   IOField "I/O field_9" at 378,310 size 30x20; FormatPattern 99
      ProcessValue <- "Motors_DB_M3_Wait_On_Now"
   IOField "I/O field_10" at 378,333 size 30x20; FormatPattern 99
      ProcessValue <- "Motors_DB_M3_Wait_Off_Now"
   IOField "I/O field_11" at 313,383 size 98x20; FormatPattern 9999999999
      ProcessValue <- "Motors_DB_M3_Res_h"
   Button "Button_45" at 213,384 size 90x20; TextOff 'Force'
      on Click: InvertBit("Motors_DB_M3_CMD_Force")
      Appearance <- "Motors_DB_M3_CMD_Force"

screen "Trans" 800x480, template "Main"
   TextField "Text field_2" at 210,15 size 67x22; Text 'Датчик:'
   TextField "Text field_4" at 273,15 size 94x22; Text 'Мутность 1'
   TextField "Text field_7" at 390,18 size 43x22; Text 'вход'
   TextField "Text field_8" at 390,43 size 56x22; Text 'выход'
   IOField "I/O field_1" at 452,19 size 102x26; FormatPattern s99999.99
      ProcessValue <- "AIx_DB_Trans_1_Converter_Min_In"
   IOField "I/O field_2" at 452,41 size 102x26; FormatPattern s99999.99
      ProcessValue <- "AIx_DB_Trans_1_Converter_Min_Out"
   IOField "I/O field_3" at 551,19 size 102x26; FormatPattern s99999.99
      ProcessValue <- "AIx_DB_Trans_1_Converter_Max_In"
   IOField "I/O field_4" at 551,41 size 102x26; FormatPattern s99999.99
      ProcessValue <- "AIx_DB_Trans_1_Converter_Max_Out"
   TextField "Text field_9" at 389,68 size 101x22; Text 'Фильтрация'
   TextField "Text field_10" at 390,96 size 36x22; Text 'RTD'
   Button "Button_7" at 489,71 size 20x20; TextOff 'Text'; PictureList "ok"
      on Click: InvertBit("AIx_DB_Trans_1_Use_Filter")
      ProcessValue <- "AIx_DB_Trans_1_Use_Filter"
   Button "Button_8" at 489,96 size 20x20; TextOff 'Text'; PictureList "ok"
      on Click: InvertBit("AIx_DB_Trans_1_Use_RTD")
      ProcessValue <- "AIx_DB_Trans_1_Use_RTD"
   IOField "I/O field_5" at 516,68 size 65x25; FormatPattern 999
      ProcessValue <- "AIx_DB_Trans_1_Filter_SP"
   IOField "I/O field_6" at 516,93 size 65x25; FormatPattern 999
      ProcessValue <- "AIx_DB_Trans_1_RTD_c"
   TextField "Text field_11" at 210,36 size 79x22; Text 'Поправка'
   IOField "I/O field_7" at 293,36 size 78x23; FormatPattern s999.9
      ProcessValue <- "AIx_DB_Trans_1_Calibration"
   Button "Button_9" at 396,176 size 248x28; TextOff 'Use'
      on Click: InvertBit("AIx_DB_Trans_1_CMD_Start_A")
      Appearance <- "AIx_DB_Trans_1_CMD_Start_A"
   Button "Button_10" at 213,66 size 68x28; TextOff 'Hand'
      on Click: InvertBit("AIx_DB_Trans_1_CMD_Hand")
      Appearance <- "AIx_DB_Trans_1_CMD_Hand"
   IOField "I/O field_8" at 293,66 size 78x28; FormatPattern s9999.9
      ProcessValue <- "AIx_DB_Trans_1_Result"
   TextField "Text field_12" at 436,123 size 27x22; Text 'NC'
   TextField "Text field_13" at 437,143 size 25x22; Text 'SC'
   TextField "Text field_14" at 210,125 size 27x22; Text 'HH'
   TextField "Text field_15" at 216,145 size 16x22; Text 'H'
   TextField "Text field_16" at 217,165 size 14x22; Text 'L'
   TextField "Text field_17" at 212,186 size 23x22; Text 'LL'
   IOField "I/O field_11" at 472,123 size 58x21; FormatPattern s99999
      ProcessValue <- "AIx_DB_Trans_1_SP_NC"
   IOField "I/O field_12" at 472,143 size 58x21; FormatPattern s99999
      ProcessValue <- "AIx_DB_Trans_1_SP_SC"
   IOField "I/O field_13" at 246,125 size 58x21; FormatPattern 99999
      ProcessValue <- "AIx_DB_Trans_1_SP_HH"
   IOField "I/O field_14" at 246,145 size 58x21; FormatPattern 99999
      ProcessValue <- "AIx_DB_Trans_1_SP_H"
   IOField "I/O field_15" at 246,165 size 58x21; FormatPattern s99999
      ProcessValue <- "AIx_DB_Trans_1_SP_L"
   IOField "I/O field_16" at 246,185 size 58x21; FormatPattern s99999
      ProcessValue <- "AIx_DB_Trans_1_SP_LL"
   IOField "I/O field_17" at 546,123 size 58x21; FormatPattern 999
      ProcessValue <- "AIx_DB_Trans_1_Timers_NC_SP"
   IOField "I/O field_18" at 546,143 size 58x21; FormatPattern 999
      ProcessValue <- "AIx_DB_Trans_1_Timers_SC_SP"
   IOField "I/O field_19" at 320,125 size 58x21; FormatPattern 999
      ProcessValue <- "AIx_DB_Trans_1_Timers_HH_SP"
   IOField "I/O field_20" at 320,145 size 58x21; FormatPattern 999
      ProcessValue <- "AIx_DB_Trans_1_Timers_H_SP"
   IOField "I/O field_21" at 320,165 size 58x21; FormatPattern 999
      ProcessValue <- "AIx_DB_Trans_1_Timers_L_SP"
   IOField "I/O field_22" at 320,185 size 58x21; FormatPattern 999
      ProcessValue <- "AIx_DB_Trans_1_Timers_LL_SP"
   IOField "I/O field_23" at 582,93 size 65x25; FormatPattern s99999
      ProcessValue <- "AIx_DB_Trans_1_Signal"
   TextField "Text field_18" at 210,97 size 68x22; Text 'Уставка'
   TextField "Text field_19" at 299,97 size 79x22; Text 'Время (с)'
   TextField "Text field_1" at 214,248 size 67x22; Text 'Датчик:'
   TextField "Text field_3" at 277,248 size 94x22; Text 'Мутность 2'
   TextField "Text field_5" at 394,251 size 43x22; Text 'вход'
   TextField "Text field_6" at 394,276 size 56x22; Text 'выход'
   IOField "I/O field_9" at 456,252 size 102x26; FormatPattern s99999.99
      ProcessValue <- "AIx_DB_Trans_2_Converter_Min_In"
   IOField "I/O field_10" at 456,274 size 102x26; FormatPattern s99999.99
      ProcessValue <- "AIx_DB_Trans_2_Converter_Min_Out"
   IOField "I/O field_24" at 555,252 size 102x26; FormatPattern s99999.99
      ProcessValue <- "AIx_DB_Trans_2_Converter_Max_In"
   IOField "I/O field_25" at 555,274 size 102x26; FormatPattern s99999.99
      ProcessValue <- "AIx_DB_Trans_2_Converter_Max_Out"
   TextField "Text field_20" at 393,301 size 101x22; Text 'Фильтрация'
   TextField "Text field_21" at 394,329 size 36x22; Text 'RTD'
   Button "Button_11" at 493,304 size 20x20; TextOff 'Text'; PictureList "ok"
      on Click: InvertBit("AIx_DB_Trans_2_Use_Filter")
      ProcessValue <- "AIx_DB_Trans_2_Use_Filter"
   Button "Button_12" at 493,329 size 20x20; TextOff 'Text'; PictureList "ok"
      on Click: InvertBit("AIx_DB_Trans_2_Use_RTD")
      ProcessValue <- "AIx_DB_Trans_2_Use_RTD"
   IOField "I/O field_26" at 520,301 size 65x25; FormatPattern 999
      ProcessValue <- "AIx_DB_Trans_2_Filter_SP"
   IOField "I/O field_27" at 520,326 size 65x25; FormatPattern 999
      ProcessValue <- "AIx_DB_Trans_2_RTD_c"
   TextField "Text field_22" at 214,269 size 79x22; Text 'Поправка'
   IOField "I/O field_28" at 297,269 size 78x23; FormatPattern s999.9
      ProcessValue <- "AIx_DB_Trans_2_Calibration"
   Button "Button_13" at 400,409 size 248x28; TextOff 'Use'
      on Click: InvertBit("AIx_DB_Trans_2_CMD_Start_A")
      Appearance <- "AIx_DB_Trans_2_CMD_Start_A"
   Button "Button_14" at 217,299 size 68x28; TextOff 'Hand'
      on Click: InvertBit("AIx_DB_Trans_2_CMD_Hand")
      Appearance <- "AIx_DB_Trans_2_CMD_Hand"
   IOField "I/O field_29" at 297,299 size 78x28; FormatPattern s9999.9
      ProcessValue <- "AIx_DB_Trans_2_Result"
   TextField "Text field_23" at 440,356 size 27x22; Text 'NC'
   TextField "Text field_24" at 441,376 size 25x22; Text 'SC'
   TextField "Text field_25" at 214,358 size 27x22; Text 'HH'
   TextField "Text field_26" at 220,378 size 16x22; Text 'H'
   TextField "Text field_27" at 221,398 size 14x22; Text 'L'
   TextField "Text field_28" at 216,419 size 23x22; Text 'LL'
   IOField "I/O field_30" at 476,356 size 58x21; FormatPattern s99999
      ProcessValue <- "AIx_DB_Trans_2_SP_NC"
   IOField "I/O field_31" at 476,376 size 58x21; FormatPattern s99999
      ProcessValue <- "AIx_DB_Trans_2_SP_SC"
   IOField "I/O field_32" at 250,358 size 58x21; FormatPattern 99999
      ProcessValue <- "AIx_DB_Trans_2_SP_HH"
   IOField "I/O field_33" at 250,378 size 58x21; FormatPattern 99999
      ProcessValue <- "AIx_DB_Trans_2_SP_H"
   IOField "I/O field_34" at 250,398 size 58x21; FormatPattern s99999
      ProcessValue <- "AIx_DB_Trans_2_SP_L"
   IOField "I/O field_35" at 250,418 size 58x21; FormatPattern s99999
      ProcessValue <- "AIx_DB_Trans_2_SP_LL"
   IOField "I/O field_36" at 550,356 size 58x21; FormatPattern 999
      ProcessValue <- "AIx_DB_Trans_2_Timers_NC_SP"
   IOField "I/O field_37" at 550,376 size 58x21; FormatPattern 999
      ProcessValue <- "AIx_DB_Trans_2_Timers_SC_SP"
   IOField "I/O field_38" at 324,358 size 58x21; FormatPattern 999
      ProcessValue <- "AIx_DB_Trans_2_Timers_HH_SP"
   IOField "I/O field_39" at 324,378 size 58x21; FormatPattern 999
      ProcessValue <- "AIx_DB_Trans_2_Timers_H_SP"
   IOField "I/O field_40" at 324,398 size 58x21; FormatPattern 999
      ProcessValue <- "AIx_DB_Trans_2_Timers_L_SP"
   IOField "I/O field_41" at 324,418 size 58x21; FormatPattern 999
      ProcessValue <- "AIx_DB_Trans_2_Timers_LL_SP"
   IOField "I/O field_42" at 586,326 size 65x25; FormatPattern s99999
      ProcessValue <- "AIx_DB_Trans_2_Signal"
   TextField "Text field_29" at 214,330 size 68x22; Text 'Уставка'
   TextField "Text field_30" at 303,330 size 79x22; Text 'Время (с)'
   Button "Button_1" at 7,5 size 96x32; TextOff 'Насосы'; Authorization "Admin"
      on Release: ActivateScreen("Dos", 0); SetTag("settings", 1)
      Appearance <- "settings"
   Button "Button_2" at 7,52 size 96x32; TextOff 'Расход'; Authorization "Admin"
      on Release: ActivateScreen("Flow", 0); SetTag("settings", 2)
      Appearance <- "settings"
   Button "Button_3" at 7,99 size 96x32; TextOff 'Мутность'; Authorization "Admin"
      on Release: ActivateScreen("Trans", 0); SetTag("settings", 3)
      Appearance <- "settings"
   Button "Button_5" at 7,146 size 96x32; TextOff 'DI'; Authorization "Admin"
      on Release: ActivateScreen("DI", 0); SetTag("settings", 4)
      Appearance <- "settings"
   Button "Button_6" at 7,193 size 96x32; TextOff 'DO'; Authorization "Admin"
      on Release: ActivateScreen("DO", 0); SetTag("settings", 5)
      Appearance <- "settings"

screen "Flow" 800x480, template "Main"
   Button "Button_1" at 7,5 size 96x32; TextOff 'Насосы'; Authorization "Admin"
      on Release: ActivateScreen("Dos", 0); SetTag("settings", 1)
      Appearance <- "settings"
   Button "Button_2" at 7,52 size 96x32; TextOff 'Расход'; Authorization "Admin"
      on Release: ActivateScreen("Flow", 0); SetTag("settings", 2)
      Appearance <- "settings"
   Button "Button_3" at 7,99 size 96x32; TextOff 'Мутность'; Authorization "Admin"
      on Release: ActivateScreen("Trans", 0); SetTag("settings", 3)
      Appearance <- "settings"
   Button "Button_5" at 7,146 size 96x32; TextOff 'DI'; Authorization "Admin"
      on Release: ActivateScreen("DI", 0); SetTag("settings", 4)
      Appearance <- "settings"
   Button "Button_6" at 7,193 size 96x32; TextOff 'DO'; Authorization "Admin"
      on Release: ActivateScreen("DO", 0); SetTag("settings", 5)
      Appearance <- "settings"
   TextField "Text field_2" at 210,15 size 67x22; Text 'Датчик:'
   TextField "Text field_4" at 273,15 size 113x22; Text 'Расходомер 1'
   TextField "Text field_7" at 390,18 size 43x22; Text 'вход'
   TextField "Text field_8" at 390,43 size 56x22; Text 'выход'
   IOField "I/O field_1" at 452,19 size 102x26; FormatPattern s99999.99
      ProcessValue <- "AIx_DB_Flow_1_Converter_Min_In"
   IOField "I/O field_2" at 452,41 size 102x26; FormatPattern s99999.99
      ProcessValue <- "AIx_DB_Flow_1_Converter_Min_Out"
   IOField "I/O field_3" at 551,19 size 102x26; FormatPattern s99999.99
      ProcessValue <- "AIx_DB_Flow_1_Converter_Max_In"
   IOField "I/O field_4" at 551,41 size 102x26; FormatPattern s99999.99
      ProcessValue <- "AIx_DB_Flow_1_Converter_Max_Out"
   TextField "Text field_9" at 389,68 size 101x22; Text 'Фильтрация'
   TextField "Text field_10" at 390,96 size 36x22; Text 'RTD'
   Button "Button_7" at 489,71 size 20x20; TextOff 'Text'; PictureList "ok"
      on Click: InvertBit("AIx_DB_Flow_1_Use_Filter")
      ProcessValue <- "AIx_DB_Flow_1_Use_Filter"
   Button "Button_8" at 489,96 size 20x20; TextOff 'Text'; PictureList "ok"
      on Click: InvertBit("AIx_DB_Flow_1_Use_RTD")
      ProcessValue <- "AIx_DB_Flow_1_Use_RTD"
   IOField "I/O field_5" at 516,68 size 65x25; FormatPattern 999
      ProcessValue <- "AIx_DB_Flow_1_Filter_SP"
   IOField "I/O field_6" at 516,93 size 65x25; FormatPattern 999
      ProcessValue <- "AIx_DB_Flow_1_RTD_c"
   TextField "Text field_11" at 210,36 size 79x22; Text 'Поправка'
   IOField "I/O field_7" at 293,36 size 78x23; FormatPattern s999.9
      ProcessValue <- "AIx_DB_Flow_1_Calibration"
   Button "Button_9" at 396,176 size 248x28; TextOff 'Use'
      on Click: InvertBit("AIx_DB_Flow_1_CMD_Start_A")
      Appearance <- "AIx_DB_Flow_1_CMD_Start_A"
   Button "Button_10" at 213,66 size 68x28; TextOff 'Hand'
      on Click: InvertBit("AIx_DB_Flow_1_CMD_Hand")
      Appearance <- "AIx_DB_Flow_1_CMD_Hand"
   IOField "I/O field_8" at 293,66 size 78x28; FormatPattern s9999.9
      ProcessValue <- "AIx_DB_Flow_1_Result"
   TextField "Text field_12" at 436,123 size 27x22; Text 'NC'
   TextField "Text field_13" at 437,143 size 25x22; Text 'SC'
   TextField "Text field_14" at 210,125 size 27x22; Text 'HH'
   TextField "Text field_15" at 216,145 size 16x22; Text 'H'
   TextField "Text field_16" at 217,165 size 14x22; Text 'L'
   TextField "Text field_17" at 212,186 size 23x22; Text 'LL'
   IOField "I/O field_11" at 472,123 size 58x21; FormatPattern s99999
      ProcessValue <- "AIx_DB_Flow_1_SP_NC"
   IOField "I/O field_12" at 472,143 size 58x21; FormatPattern s99999
      ProcessValue <- "AIx_DB_Flow_1_SP_SC"
   IOField "I/O field_13" at 246,125 size 58x21; FormatPattern 99999
      ProcessValue <- "AIx_DB_Flow_1_SP_HH"
   IOField "I/O field_14" at 246,145 size 58x21; FormatPattern 99999
      ProcessValue <- "AIx_DB_Flow_1_SP_H"
   IOField "I/O field_15" at 246,165 size 58x21; FormatPattern s99999
      ProcessValue <- "AIx_DB_Flow_1_SP_L"
   IOField "I/O field_16" at 246,185 size 58x21; FormatPattern s99999
      ProcessValue <- "AIx_DB_Flow_1_SP_LL"
   IOField "I/O field_17" at 546,123 size 58x21; FormatPattern 999
      ProcessValue <- "AIx_DB_Flow_1_Timers_NC_SP"
   IOField "I/O field_18" at 546,143 size 58x21; FormatPattern 999
      ProcessValue <- "AIx_DB_Flow_1_Timers_SC_SP"
   IOField "I/O field_19" at 320,125 size 58x21; FormatPattern 999
      ProcessValue <- "AIx_DB_Flow_1_Timers_HH_SP"
   IOField "I/O field_20" at 320,145 size 58x21; FormatPattern 999
      ProcessValue <- "AIx_DB_Flow_1_Timers_H_SP"
   IOField "I/O field_21" at 320,165 size 58x21; FormatPattern 999
      ProcessValue <- "AIx_DB_Flow_1_Timers_L_SP"
   IOField "I/O field_22" at 320,185 size 58x21; FormatPattern 999
      ProcessValue <- "AIx_DB_Flow_1_Timers_LL_SP"
   IOField "I/O field_23" at 582,93 size 65x25; FormatPattern s99999
      ProcessValue <- "AIx_DB_Flow_1_Signal"
   TextField "Text field_18" at 210,97 size 68x22; Text 'Уставка'
   TextField "Text field_19" at 299,97 size 79x22; Text 'Время (с)'
   TextField "Text field_1" at 214,248 size 67x22; Text 'Датчик:'
   TextField "Text field_3" at 277,248 size 113x22; Text 'Расходомер 2'
   TextField "Text field_5" at 394,251 size 43x22; Text 'вход'
   TextField "Text field_6" at 394,276 size 56x22; Text 'выход'
   IOField "I/O field_9" at 456,252 size 102x26; FormatPattern s99999.99
      ProcessValue <- "AIx_DB_Flow_2_Converter_Min_In"
   IOField "I/O field_10" at 456,274 size 102x26; FormatPattern s99999.99
      ProcessValue <- "AIx_DB_Flow_2_Converter_Min_Out"
   IOField "I/O field_24" at 555,252 size 102x26; FormatPattern s99999.99
      ProcessValue <- "AIx_DB_Flow_2_Converter_Max_In"
   IOField "I/O field_25" at 555,274 size 102x26; FormatPattern s99999.99
      ProcessValue <- "AIx_DB_Flow_2_Converter_Max_Out"
   TextField "Text field_20" at 393,301 size 101x22; Text 'Фильтрация'
   TextField "Text field_21" at 394,329 size 36x22; Text 'RTD'
   Button "Button_11" at 493,304 size 20x20; TextOff 'Text'; PictureList "ok"
      on Click: InvertBit("AIx_DB_Flow_2_Use_Filter")
      ProcessValue <- "AIx_DB_Flow_2_Use_Filter"
   Button "Button_12" at 493,329 size 20x20; TextOff 'Text'; PictureList "ok"
      on Click: InvertBit("AIx_DB_Flow_2_Use_RTD")
      ProcessValue <- "AIx_DB_Flow_2_Use_RTD"
   IOField "I/O field_26" at 520,301 size 65x25; FormatPattern 999
      ProcessValue <- "AIx_DB_Flow_2_Filter_SP"
   IOField "I/O field_27" at 520,326 size 65x25; FormatPattern 999
      ProcessValue <- "AIx_DB_Flow_2_RTD_c"
   TextField "Text field_22" at 214,269 size 79x22; Text 'Поправка'
   IOField "I/O field_28" at 297,269 size 78x23; FormatPattern s999.9
      ProcessValue <- "AIx_DB_Flow_2_Calibration"
   Button "Button_13" at 400,409 size 248x28; TextOff 'Use'
      on Click: InvertBit("AIx_DB_Flow_2_CMD_Start_A")
      Appearance <- "AIx_DB_Flow_2_CMD_Start_A"
   Button "Button_14" at 217,299 size 68x28; TextOff 'Hand'
      on Click: InvertBit("AIx_DB_Flow_2_CMD_Hand")
      Appearance <- "AIx_DB_Flow_2_CMD_Hand"
   IOField "I/O field_29" at 297,299 size 78x28; FormatPattern s9999.9
      ProcessValue <- "AIx_DB_Flow_2_Result"
   TextField "Text field_23" at 440,356 size 27x22; Text 'NC'
   TextField "Text field_24" at 441,376 size 25x22; Text 'SC'
   TextField "Text field_25" at 214,358 size 27x22; Text 'HH'
   TextField "Text field_26" at 220,378 size 16x22; Text 'H'
   TextField "Text field_27" at 221,398 size 14x22; Text 'L'
   TextField "Text field_28" at 216,419 size 23x22; Text 'LL'
   IOField "I/O field_30" at 476,356 size 58x21; FormatPattern s99999
      ProcessValue <- "AIx_DB_Flow_2_SP_NC"
   IOField "I/O field_31" at 476,376 size 58x21; FormatPattern s99999
      ProcessValue <- "AIx_DB_Flow_2_SP_SC"
   IOField "I/O field_32" at 250,358 size 58x21; FormatPattern 99999
      ProcessValue <- "AIx_DB_Flow_2_SP_HH"
   IOField "I/O field_33" at 250,378 size 58x21; FormatPattern 99999
      ProcessValue <- "AIx_DB_Flow_2_SP_H"
   IOField "I/O field_34" at 250,398 size 58x21; FormatPattern s99999
      ProcessValue <- "AIx_DB_Flow_2_SP_L"
   IOField "I/O field_35" at 250,418 size 58x21; FormatPattern s99999
      ProcessValue <- "AIx_DB_Flow_2_SP_LL"
   IOField "I/O field_36" at 550,356 size 58x21; FormatPattern 999
      ProcessValue <- "AIx_DB_Flow_2_Timers_NC_SP"
   IOField "I/O field_37" at 550,376 size 58x21; FormatPattern 999
      ProcessValue <- "AIx_DB_Flow_2_Timers_SC_SP"
   IOField "I/O field_38" at 324,358 size 58x21; FormatPattern 999
      ProcessValue <- "AIx_DB_Flow_2_Timers_HH_SP"
   IOField "I/O field_39" at 324,378 size 58x21; FormatPattern 999
      ProcessValue <- "AIx_DB_Flow_2_Timers_H_SP"
   IOField "I/O field_40" at 324,398 size 58x21; FormatPattern 999
      ProcessValue <- "AIx_DB_Flow_2_Timers_L_SP"
   IOField "I/O field_41" at 324,418 size 58x21; FormatPattern 999
      ProcessValue <- "AIx_DB_Flow_2_Timers_LL_SP"
   IOField "I/O field_42" at 586,326 size 65x25; FormatPattern s99999
      ProcessValue <- "AIx_DB_Flow_2_Signal"
   TextField "Text field_29" at 214,330 size 68x22; Text 'Уставка'
   TextField "Text field_30" at 303,330 size 79x22; Text 'Время (с)'

screen "DI" 800x480, template "Main"
   Group "Group" at 127,7 size 283x51; TextList "Hand"
   Group "Group_1" at 127,66 size 283x51; TextList "Hand"
   Group "Group_2" at 127,125 size 283x51; TextList "Hand"
   Group "Group_3" at 127,184 size 283x51; TextList "Hand"
   Group "Group_4" at 127,244 size 283x51; TextList "Hand"
   Group "Group_5" at 127,303 size 283x51; TextList "Hand"
   Group "Group_6" at 127,362 size 283x51; TextList "Hand"
   Group "Group_7" at 127,422 size 283x51; TextList "Hand"
   Group "Group_8" at 433,7 size 283x51; TextList "Hand"
   Group "Group_9" at 433,66 size 283x51; TextList "Hand"
   Button "Button_1" at 7,5 size 96x32; TextOff 'Насосы'; Authorization "Admin"
      on Release: ActivateScreen("Dos", 0); SetTag("settings", 1)
      Appearance <- "settings"
   Button "Button_2" at 7,52 size 96x32; TextOff 'Расход'; Authorization "Admin"
      on Release: ActivateScreen("Flow", 0); SetTag("settings", 2)
      Appearance <- "settings"
   Button "Button_3" at 7,99 size 96x32; TextOff 'Мутность'; Authorization "Admin"
      on Release: ActivateScreen("Trans", 0); SetTag("settings", 3)
      Appearance <- "settings"
   Button "Button_5" at 7,146 size 96x32; TextOff 'DI'; Authorization "Admin"
      on Release: ActivateScreen("DI", 0); SetTag("settings", 4)
      Appearance <- "settings"
   Button "Button_6" at 7,193 size 96x32; TextOff 'DO'; Authorization "Admin"
      on Release: ActivateScreen("DO", 0); SetTag("settings", 5)
      Appearance <- "settings"
   TextField "Text field_1" at 131,10 size 45x22; Text 'I 0.0'
   TextField "Text field_2" at 176,10 size 120x22; Text 'M1 Готовность'
   Circle "Circle_1" at 131,33 size 22x22
      Appearance <- "DIx_DB_M1_QF_Input"
   Circle "Circle_2" at 154,33 size 22x22
      Appearance <- "DIx_DB_M1_QF_Signal"
   Button "Button_7" at 298,11 size 59x44; TextOff 'Авто'; TextList "Hand"
      on Click: InvertBit("DIx_DB_M1_QF_Hand")
      Appearance <- "DIx_DB_M1_QF_Hand"
      ProcessValue <- "DIx_DB_M1_QF_Hand"
   Button "Button_8" at 240,33 size 49x22; TextOff 'Выкл'
      on Click: ResetBit("DIx_DB_M1_QF_Start_M")
   Button "Button_12" at 184,33 size 47x22; TextOff 'Вкл'
      on Click: SetBit("DIx_DB_M1_QF_Start_M")
      Appearance <- "DIx_DB_M1_QF_Start_M"
   IOField "I/O field_6" at 360,33 size 23x22; FormatPattern 99
      ProcessValue <- "DIx_DB_M1_QF_Filter_On_SP"
   IOField "I/O field_7" at 383,33 size 23x22; FormatPattern 99
      ProcessValue <- "DIx_DB_M1_QF_Filter_Off_SP"
   Button "Button_9" at 360,10 size 46x20; TextOff 'Inv'
      on Click: InvertBit("DIx_DB_M1_QF_Inverse")
      Appearance <- "DIx_DB_M1_QF_Inverse"
   TextField "Text field_3" at 131,69 size 45x22; Text 'I 0.1'
   TextField "Text field_4" at 176,69 size 120x22; Text 'М2 Готовность'
   Circle "Circle_3" at 131,92 size 22x22
      Appearance <- "DIx_DB_M2_QF_Input"
   Circle "Circle_4" at 154,92 size 22x22
      Appearance <- "DIx_DB_M2_QF_Signal"
   Button "Button_10" at 298,70 size 59x44; TextOff 'Авто'; TextList "Hand"
      on Click: InvertBit("DIx_DB_M2_QF_Hand")
      Appearance <- "DIx_DB_M2_QF_Hand"
      ProcessValue <- "DIx_DB_M2_QF_Hand"
   Button "Button_11" at 240,92 size 49x22; TextOff 'Выкл'
      on Click: ResetBit("DIx_DB_M2_QF_Start_M")
   Button "Button_13" at 184,92 size 47x22; TextOff 'Вкл'
      on Click: SetBit("DIx_DB_M2_QF_Start_M")
      Appearance <- "DIx_DB_M2_QF_Start_M"
   IOField "I/O field_1" at 360,92 size 23x22; FormatPattern 99
      ProcessValue <- "DIx_DB_M2_QF_Filter_On_SP"
   IOField "I/O field_2" at 383,92 size 23x22; FormatPattern 99
      ProcessValue <- "DIx_DB_M2_QF_Filter_Off_SP"
   Button "Button_14" at 360,69 size 46x20; TextOff 'Inv'
      on Click: InvertBit("DIx_DB_M2_QF_Inverse")
      Appearance <- "DIx_DB_M2_QF_Inverse"
   TextField "Text field_5" at 131,128 size 45x22; Text 'I 0.2'
   TextField "Text field_6" at 176,128 size 120x22; Text 'M3 Готовность'
   Circle "Circle_5" at 131,151 size 22x22
      Appearance <- "DIx_DB_M3_QF_Input"
   Circle "Circle_6" at 154,151 size 22x22
      Appearance <- "DIx_DB_M3_QF_Signal"
   Button "Button_15" at 298,129 size 59x44; TextOff 'Авто'; TextList "Hand"
      on Click: InvertBit("DIx_DB_M3_QF_Hand")
      Appearance <- "DIx_DB_M3_QF_Hand"
      ProcessValue <- "DIx_DB_M3_QF_Hand"
   Button "Button_16" at 240,151 size 49x22; TextOff 'Выкл'
      on Click: ResetBit("DIx_DB_M3_QF_Start_M")
   Button "Button_17" at 184,151 size 47x22; TextOff 'Вкл'
      on Click: SetBit("DIx_DB_M3_QF_Start_M")
      Appearance <- "DIx_DB_M3_QF_Start_M"
   IOField "I/O field_3" at 360,151 size 23x22; FormatPattern 99
      ProcessValue <- "DIx_DB_M3_QF_Filter_On_SP"
   IOField "I/O field_4" at 383,151 size 23x22; FormatPattern 99
      ProcessValue <- "DIx_DB_M3_QF_Filter_Off_SP"
   Button "Button_18" at 360,128 size 46x20; TextOff 'Inv'
      on Click: InvertBit("DIx_DB_M3_QF_Inverse")
      Appearance <- "DIx_DB_M3_QF_Inverse"
   TextField "Text field_7" at 131,187 size 45x22; Text 'I 0.3'
   TextField "Text field_8" at 176,187 size 119x22; Text 'Нагреватель 1'
   Circle "Circle_7" at 131,210 size 22x22
      Appearance <- "DIx_DB_Heat_1_Input"
   Circle "Circle_8" at 154,210 size 22x22
      Appearance <- "DIx_DB_Heat_1_Signal"
   Button "Button_19" at 298,188 size 59x44; TextOff 'Авто'; TextList "Hand"
      on Click: InvertBit("DIx_DB_Heat_1_Hand")
      Appearance <- "DIx_DB_Heat_1_Hand"
      ProcessValue <- "DIx_DB_Heat_1_Hand"
   Button "Button_20" at 240,210 size 49x22; TextOff 'Выкл'
      on Click: ResetBit("DIx_DB_Heat_1_Start_M")
   Button "Button_21" at 184,210 size 47x22; TextOff 'Вкл'
      on Click: SetBit("DIx_DB_Heat_1_Start_M")
      Appearance <- "DIx_DB_Heat_1_Start_M"
   IOField "I/O field_5" at 360,210 size 23x22; FormatPattern 99
      ProcessValue <- "DIx_DB_Heat_1_Filter_On_SP"
   IOField "I/O field_8" at 383,210 size 23x22; FormatPattern 99
      ProcessValue <- "DIx_DB_Heat_1_Filter_Off_SP"
   Button "Button_22" at 360,187 size 46x20; TextOff 'Inv'
      on Click: InvertBit("DIx_DB_Heat_1_Inverse")
      Appearance <- "DIx_DB_Heat_1_Inverse"
   TextField "Text field_9" at 131,247 size 45x22; Text 'I 0.4'
   TextField "Text field_10" at 176,247 size 119x22; Text 'Нагреватель 2'
   Circle "Circle_9" at 131,270 size 22x22
      Appearance <- "DIx_DB_Heat_2_Input"
   Circle "Circle_10" at 154,270 size 22x22
      Appearance <- "DIx_DB_Heat_2_Signal"
   Button "Button_23" at 298,248 size 59x44; TextOff 'Авто'; TextList "Hand"
      on Click: InvertBit("DIx_DB_Heat_2_Hand")
      Appearance <- "DIx_DB_Heat_2_Hand"
      ProcessValue <- "DIx_DB_Heat_2_Hand"
   Button "Button_24" at 240,270 size 49x22; TextOff 'Выкл'
      on Click: ResetBit("DIx_DB_Heat_2_Start_M")
   Button "Button_25" at 184,270 size 47x22; TextOff 'Вкл'
      on Click: SetBit("DIx_DB_Heat_2_Start_M")
      Appearance <- "DIx_DB_Heat_2_Start_M"
   IOField "I/O field_9" at 360,270 size 23x22; FormatPattern 99
      ProcessValue <- "DIx_DB_Heat_2_Filter_On_SP"
   IOField "I/O field_10" at 383,270 size 23x22; FormatPattern 99
      ProcessValue <- "DIx_DB_Heat_2_Filter_Off_SP"
   Button "Button_26" at 360,247 size 46x20; TextOff 'Inv'
      on Click: InvertBit("DIx_DB_Heat_2_Inverse")
      Appearance <- "DIx_DB_Heat_2_Inverse"
   TextField "Text field_11" at 131,306 size 45x22; Text 'I 0.5'
   TextField "Text field_12" at 176,306 size 119x22; Text 'Нагреватель 3'
   Circle "Circle_11" at 131,329 size 22x22
      Appearance <- "DIx_DB_Heat_3_Input"
   Circle "Circle_12" at 154,329 size 22x22
      Appearance <- "DIx_DB_Heat_3_Signal"
   Button "Button_27" at 298,307 size 59x44; TextOff 'Авто'; TextList "Hand"
      on Click: InvertBit("DIx_DB_Heat_3_Hand")
      Appearance <- "DIx_DB_Heat_3_Hand"
      ProcessValue <- "DIx_DB_Heat_3_Hand"
   Button "Button_28" at 240,329 size 49x22; TextOff 'Выкл'
      on Click: ResetBit("DIx_DB_Heat_3_Start_M")
   Button "Button_29" at 184,329 size 47x22; TextOff 'Вкл'
      on Click: SetBit("DIx_DB_Heat_3_Start_M")
      Appearance <- "DIx_DB_Heat_3_Start_M"
   IOField "I/O field_11" at 360,329 size 23x22; FormatPattern 99
      ProcessValue <- "DIx_DB_Heat_3_Filter_On_SP"
   IOField "I/O field_12" at 383,329 size 23x22; FormatPattern 99
      ProcessValue <- "DIx_DB_Heat_3_Filter_Off_SP"
   Button "Button_30" at 360,306 size 46x20; TextOff 'Inv'
      on Click: InvertBit("DIx_DB_Heat_3_Inverse")
      Appearance <- "DIx_DB_Heat_3_Inverse"
   TextField "Text field_13" at 131,365 size 45x22; Text 'I 0.6'
   TextField "Text field_14" at 176,365 size 119x22; Text 'Нагреватель 4'
   Circle "Circle_13" at 131,388 size 22x22
      Appearance <- "DIx_DB_Heat_4_Input"
   Circle "Circle_14" at 154,388 size 22x22
      Appearance <- "DIx_DB_Heat_4_Signal"
   Button "Button_31" at 298,366 size 59x44; TextOff 'Авто'; TextList "Hand"
      on Click: InvertBit("DIx_DB_Heat_4_Hand")
      Appearance <- "DIx_DB_Heat_4_Hand"
      ProcessValue <- "DIx_DB_Heat_4_Hand"
   Button "Button_32" at 240,388 size 49x22; TextOff 'Выкл'
      on Click: ResetBit("DIx_DB_Heat_4_Start_M")
   Button "Button_33" at 184,388 size 47x22; TextOff 'Вкл'
      on Click: SetBit("DIx_DB_Heat_4_Start_M")
      Appearance <- "DIx_DB_Heat_4_Start_M"
   IOField "I/O field_13" at 360,388 size 23x22; FormatPattern 99
      ProcessValue <- "DIx_DB_Heat_4_Filter_On_SP"
   IOField "I/O field_14" at 383,388 size 23x22; FormatPattern 99
      ProcessValue <- "DIx_DB_Heat_4_Filter_Off_SP"
   Button "Button_34" at 360,365 size 46x20; TextOff 'Inv'
      on Click: InvertBit("DIx_DB_Heat_4_Inverse")
      Appearance <- "DIx_DB_Heat_4_Inverse"
   TextField "Text field_15" at 131,425 size 45x22; Text 'I 0.7'
   TextField "Text field_16" at 176,425 size 112x22; Text 'Внешний стоп'
   Circle "Circle_15" at 131,448 size 22x22
      Appearance <- "DIx_DB_AllBlock_Input"
   Circle "Circle_16" at 154,448 size 22x22
      Appearance <- "DIx_DB_AllBlock_Signal"
   Button "Button_35" at 298,426 size 59x44; TextOff 'Авто'; TextList "Hand"
      on Click: InvertBit("DIx_DB_AllBlock_Hand")
      Appearance <- "DIx_DB_AllBlock_Hand"
      ProcessValue <- "DIx_DB_AllBlock_Hand"
   Button "Button_36" at 240,448 size 49x22; TextOff 'Выкл'
      on Click: ResetBit("DIx_DB_AllBlock_Start_M")
   Button "Button_37" at 184,448 size 47x22; TextOff 'Вкл'
      on Click: SetBit("DIx_DB_AllBlock_Start_M")
      Appearance <- "DIx_DB_AllBlock_Start_M"
   IOField "I/O field_15" at 360,448 size 23x22; FormatPattern 99
      ProcessValue <- "DIx_DB_AllBlock_Filter_On_SP"
   IOField "I/O field_16" at 383,448 size 23x22; FormatPattern 99
      ProcessValue <- "DIx_DB_AllBlock_Filter_Off_SP"
   Button "Button_38" at 360,425 size 46x20; TextOff 'Inv'
      on Click: InvertBit("DIx_DB_AllBlock_Inverse")
      Appearance <- "DIx_DB_AllBlock_Inverse"
   TextField "Text field_17" at 437,10 size 45x22; Text 'I 1.0'
   TextField "Text field_18" at 482,10 size 59x22; Text 'Весы 1'
   Circle "Circle_17" at 437,33 size 22x22
      Appearance <- "DIx_DB_Mass_1_Input"
   Circle "Circle_18" at 460,33 size 22x22
      Appearance <- "DIx_DB_Mass_1_Signal"
   Button "Button_39" at 604,11 size 59x44; TextOff 'Авто'; TextList "Hand"
      on Click: InvertBit("DIx_DB_Mass_1_Hand")
      Appearance <- "DIx_DB_Mass_1_Hand"
      ProcessValue <- "DIx_DB_Mass_1_Hand"
   Button "Button_40" at 546,33 size 49x22; TextOff 'Выкл'
      on Click: ResetBit("DIx_DB_Mass_1_Start_M")
   Button "Button_41" at 490,33 size 47x22; TextOff 'Вкл'
      on Click: SetBit("DIx_DB_Mass_1_Start_M")
      Appearance <- "DIx_DB_Mass_1_Start_M"
   IOField "I/O field_17" at 666,33 size 23x22; FormatPattern 99
      ProcessValue <- "DIx_DB_Mass_1_Filter_On_SP"
   IOField "I/O field_18" at 689,33 size 23x22; FormatPattern 99
      ProcessValue <- "DIx_DB_Mass_1_Filter_Off_SP"
   Button "Button_42" at 666,10 size 46x20; TextOff 'Inv'
      on Click: InvertBit("DIx_DB_Mass_1_Inverse")
      Appearance <- "DIx_DB_Mass_1_Inverse"
   TextField "Text field_19" at 437,69 size 45x22; Text 'I 1.1'
   TextField "Text field_20" at 482,69 size 59x22; Text 'Весы 2'
   Circle "Circle_19" at 437,92 size 22x22
      Appearance <- "DIx_DB_Mass_2_Input"
   Circle "Circle_20" at 460,92 size 22x22
      Appearance <- "DIx_DB_Mass_2_Signal"
   Button "Button_43" at 604,70 size 59x44; TextOff 'Авто'; TextList "Hand"
      on Click: InvertBit("DIx_DB_Mass_2_Hand")
      Appearance <- "DIx_DB_Mass_2_Hand"
      ProcessValue <- "DIx_DB_Mass_2_Hand"
   Button "Button_44" at 546,92 size 49x22; TextOff 'Выкл'
      on Click: ResetBit("DIx_DB_Mass_2_Start_M")
   Button "Button_45" at 490,92 size 47x22; TextOff 'Вкл'
      on Click: SetBit("DIx_DB_Mass_2_Start_M")
      Appearance <- "DIx_DB_Mass_2_Start_M"
   IOField "I/O field_19" at 666,92 size 23x22; FormatPattern 99
      ProcessValue <- "DIx_DB_Mass_2_Filter_On_SP"
   IOField "I/O field_20" at 689,92 size 23x22; FormatPattern 99
      ProcessValue <- "DIx_DB_Mass_2_Filter_Off_SP"
   Button "Button_46" at 666,69 size 46x20; TextOff 'Inv'
      on Click: InvertBit("DIx_DB_Mass_2_Inverse")
      Appearance <- "DIx_DB_Mass_2_Inverse"

screen "DO" 800x480, template "Main"
   Group "Group" at 127,7 size 283x51; TextList "Hand"
   Group "Group_1" at 127,66 size 283x51; Text 'Q 0.0'; TextList "Hand"
   Group "Group_2" at 127,125 size 283x51; Text 'Q 0.0'; TextList "Hand"
   Group "Group_3" at 127,184 size 283x51; Text 'Q 0.0'; TextList "Hand"
   Group "Group_4" at 127,244 size 283x51; Text 'Q 0.0'; TextList "Hand"
   Group "Group_5" at 127,303 size 283x51; Text 'Q 0.0'; TextList "Hand"
   Group "Group_6" at 127,362 size 283x51; Text 'Q 0.0'; TextList "Hand"
   Group "Group_7" at 127,422 size 283x51; Text 'Q 0.0'; TextList "Hand"
   Group "Group_8" at 433,7 size 283x51; Text 'Q 0.0'; TextList "Hand"
   Button "Button_1" at 7,5 size 96x32; TextOff 'Насосы'; Authorization "Admin"
      on Release: ActivateScreen("Dos", 0); SetTag("settings", 1)
      Appearance <- "settings"
   Button "Button_2" at 7,52 size 96x32; TextOff 'Расход'; Authorization "Admin"
      on Release: ActivateScreen("Flow", 0); SetTag("settings", 2)
      Appearance <- "settings"
   Button "Button_3" at 7,99 size 96x32; TextOff 'Мутность'; Authorization "Admin"
      on Release: ActivateScreen("Trans", 0); SetTag("settings", 3)
      Appearance <- "settings"
   Button "Button_5" at 7,146 size 96x32; TextOff 'DI'; Authorization "Admin"
      on Release: ActivateScreen("DI", 0); SetTag("settings", 4)
      Appearance <- "settings"
   Button "Button_6" at 7,193 size 96x32; TextOff 'DO'; Authorization "Admin"
      on Release: ActivateScreen("DO", 0); SetTag("settings", 5)
      Appearance <- "settings"
   TextField "Text field_4" at 131,10 size 45x22; Text 'Q 0.0'
   TextField "Text field_5" at 176,10 size 69x22; Text 'M1 Пуск'
   Circle "Circle_3" at 131,33 size 22x22
      Appearance <- "DOx_DB_M1_CMD_Start_A"
   Circle "Circle_4" at 154,33 size 22x22
      Appearance <- "DOx_DB_M1_CMD_Q"
   Button "Button_13" at 298,11 size 59x44; TextOff 'Авто'; TextList "Hand"
      on Click: InvertBit("DOx_DB_M1_CMD_Hand")
      Appearance <- "DOx_DB_M1_CMD_Hand"
      ProcessValue <- "DOx_DB_M1_CMD_Hand"
   Button "Button_14" at 240,33 size 49x22; TextOff 'Выкл'
      on Click: ResetBit("DOx_DB_M1_CMD_Start_M")
   Button "Button_15" at 184,33 size 47x22; TextOff 'Вкл'
      on Click: SetBit("DOx_DB_M1_CMD_Start_M")
      Appearance <- "DOx_DB_M1_CMD_Start_M"
   Button "Button_16" at 360,10 size 46x20; TextOff 'Inv'
      on Click: InvertBit("DOx_DB_M1_CMD_Inverse")
      Appearance <- "DOx_DB_M1_CMD_Inverse"
   Button "Button_17" at 360,35 size 46x20; TextOff 'Sim'
      on Click: InvertBit("DOx_DB_M1_CMD_Simulation")
      Appearance <- "DOx_DB_M1_CMD_Simulation"
   TextField "Text field_1" at 131,69 size 45x22; Text 'Q 0.1'
   TextField "Text field_2" at 176,69 size 69x22; Text 'M2 Пуск'
   Circle "Circle_1" at 131,92 size 22x22
      Appearance <- "DOx_DB_M2_CMD_Start_A"
   Circle "Circle_2" at 154,92 size 22x22
      Appearance <- "DOx_DB_M2_CMD_Q"
   Button "Button_7" at 298,70 size 59x44; TextOff 'Авто'; TextList "Hand"
      on Click: InvertBit("DOx_DB_M2_CMD_Hand")
      Appearance <- "DOx_DB_M2_CMD_Hand"
      ProcessValue <- "DOx_DB_M2_CMD_Hand"
   Button "Button_8" at 240,92 size 49x22; TextOff 'Выкл'
      on Click: ResetBit("DOx_DB_M2_CMD_Start_M")
   Button "Button_9" at 184,92 size 47x22; TextOff 'Вкл'
      on Click: SetBit("DOx_DB_M2_CMD_Start_M")
      Appearance <- "DOx_DB_M2_CMD_Start_M"
   Button "Button_10" at 360,69 size 46x20; TextOff 'Inv'
      on Click: InvertBit("DOx_DB_M2_CMD_Inverse")
      Appearance <- "DOx_DB_M2_CMD_Inverse"
   Button "Button_11" at 360,94 size 46x20; TextOff 'Sim'
      on Click: InvertBit("DOx_DB_M2_CMD_Simulation")
      Appearance <- "DOx_DB_M2_CMD_Simulation"
   TextField "Text field_3" at 131,128 size 45x22; Text 'Q 0.2'
   TextField "Text field_6" at 176,128 size 69x22; Text 'M3 Пуск'
   Circle "Circle_5" at 131,151 size 22x22
      Appearance <- "DOx_DB_M3_CMD_Start_A"
   Circle "Circle_6" at 154,151 size 22x22
      Appearance <- "DOx_DB_M3_CMD_Q"
   Button "Button_12" at 298,129 size 59x44; TextOff 'Авто'; TextList "Hand"
      on Click: InvertBit("DOx_DB_M3_CMD_Hand")
      Appearance <- "DOx_DB_M3_CMD_Hand"
      ProcessValue <- "DOx_DB_M3_CMD_Hand"
   Button "Button_18" at 240,151 size 49x22; TextOff 'Выкл'
      on Click: ResetBit("DOx_DB_M3_CMD_Start_M")
   Button "Button_19" at 184,151 size 47x22; TextOff 'Вкл'
      on Click: SetBit("DOx_DB_M3_CMD_Start_M")
      Appearance <- "DOx_DB_M3_CMD_Start_M"
   Button "Button_20" at 360,128 size 46x20; TextOff 'Inv'
      on Click: InvertBit("DOx_DB_M3_CMD_Inverse")
      Appearance <- "DOx_DB_M3_CMD_Inverse"
   Button "Button_21" at 360,153 size 46x20; TextOff 'Sim'
      on Click: InvertBit("DOx_DB_M3_CMD_Simulation")
      Appearance <- "DOx_DB_M3_CMD_Simulation"
   TextField "Text field_7" at 131,187 size 45x22; Text 'Q 0.3'
   TextField "Text field_8" at 176,187 size 107x22; Text 'LED Авария 1'
   Circle "Circle_7" at 131,210 size 22x22
      Appearance <- "DOx_DB_LED_Error_1_Start_A"
   Circle "Circle_8" at 154,210 size 22x22
      Appearance <- "DOx_DB_LED_Error_1_Q"
   Button "Button_22" at 298,188 size 59x44; TextOff 'Авто'; TextList "Hand"
      on Click: InvertBit("DOx_DB_LED_Error_1_Hand")
      Appearance <- "DOx_DB_LED_Error_1_Hand"
      ProcessValue <- "DOx_DB_LED_Error_1_Hand"
   Button "Button_23" at 240,210 size 49x22; TextOff 'Выкл'
      on Click: ResetBit("DOx_DB_LED_Error_1_Start_M")
   Button "Button_24" at 184,210 size 47x22; TextOff 'Вкл'
      on Click: SetBit("DOx_DB_LED_Error_1_Start_M")
      Appearance <- "DOx_DB_LED_Error_1_Start_M"
   Button "Button_25" at 360,187 size 46x20; TextOff 'Inv'
      on Click: InvertBit("DOx_DB_LED_Error_1_Inverse")
      Appearance <- "DOx_DB_LED_Error_1_Inverse"
   Button "Button_26" at 360,212 size 46x20; TextOff 'Sim'
      on Click: InvertBit("DOx_DB_LED_Error_1_Simulation")
      Appearance <- "DOx_DB_LED_Error_1_Simulation"
   TextField "Text field_9" at 131,247 size 45x22; Text 'Q 0.4'
   TextField "Text field_10" at 176,247 size 107x22; Text 'LED Авария 2'
   Circle "Circle_9" at 131,270 size 22x22
      Appearance <- "DOx_DB_LED_Error_2_Start_A"
   Circle "Circle_10" at 154,270 size 22x22
      Appearance <- "DOx_DB_LED_Error_2_Q"
   Button "Button_27" at 298,248 size 59x44; TextOff 'Авто'; TextList "Hand"
      on Click: InvertBit("DOx_DB_LED_Error_2_Hand")
      Appearance <- "DOx_DB_LED_Error_2_Hand"
      ProcessValue <- "DOx_DB_LED_Error_2_Hand"
   Button "Button_28" at 240,270 size 49x22; TextOff 'Выкл'
      on Click: ResetBit("DOx_DB_LED_Error_2_Start_M")
   Button "Button_29" at 184,270 size 47x22; TextOff 'Вкл'
      on Click: SetBit("DOx_DB_LED_Error_2_Start_M")
      Appearance <- "DOx_DB_LED_Error_2_Start_M"
   Button "Button_30" at 360,247 size 46x20; TextOff 'Inv'
      on Click: InvertBit("DOx_DB_LED_Error_2_Inverse")
      Appearance <- "DOx_DB_LED_Error_2_Inverse"
   Button "Button_31" at 360,272 size 46x20; TextOff 'Sim'
      on Click: InvertBit("DOx_DB_LED_Error_2_Simulation")
      Appearance <- "DOx_DB_LED_Error_2_Simulation"
   TextField "Text field_11" at 131,306 size 45x22; Text 'Q 0.5'
   TextField "Text field_12" at 176,306 size 93x22; Text 'LED Авария'
   Circle "Circle_11" at 131,329 size 22x22
      Appearance <- "DOx_DB_LED_Alarm_Start_A"
   Circle "Circle_12" at 154,329 size 22x22
      Appearance <- "DOx_DB_LED_Alarm_Q"
   Button "Button_32" at 298,307 size 59x44; TextOff 'Авто'; TextList "Hand"
      on Click: InvertBit("DOx_DB_LED_Alarm_Hand")
      Appearance <- "DOx_DB_LED_Alarm_Hand"
      ProcessValue <- "DOx_DB_LED_Alarm_Hand"
   Button "Button_33" at 240,329 size 49x22; TextOff 'Выкл'
      on Click: ResetBit("DOx_DB_LED_Alarm_Start_M")
   Button "Button_34" at 184,329 size 47x22; TextOff 'Вкл'
      on Click: SetBit("DOx_DB_LED_Alarm_Start_M")
      Appearance <- "DOx_DB_LED_Alarm_Start_M"
   Button "Button_35" at 360,306 size 46x20; TextOff 'Inv'
      on Click: InvertBit("DOx_DB_LED_Alarm_Inverse")
      Appearance <- "DOx_DB_LED_Alarm_Inverse"
   Button "Button_36" at 360,331 size 46x20; TextOff 'Sim'
      on Click: InvertBit("DOx_DB_LED_Alarm_Simulation")
      Appearance <- "DOx_DB_LED_Alarm_Simulation"
   TextField "Text field_13" at 131,365 size 45x22; Text 'Q 0.6'
   TextField "Text field_14" at 176,365 size 120x22; Text 'LED М1 Авария'
   Circle "Circle_13" at 131,388 size 22x22
      Appearance <- "DOx_DB_LED_M1_Alarm_Start_A"
   Circle "Circle_14" at 154,388 size 22x22
      Appearance <- "DOx_DB_LED_M1_Alarm_Q"
   Button "Button_37" at 298,366 size 59x44; TextOff 'Авто'; TextList "Hand"
      on Click: InvertBit("DOx_DB_LED_M1_Alarm_Hand")
      Appearance <- "DOx_DB_LED_M1_Alarm_Hand"
      ProcessValue <- "DOx_DB_LED_M1_Alarm_Hand"
   Button "Button_38" at 240,388 size 49x22; TextOff 'Выкл'
      on Click: ResetBit("DOx_DB_LED_M1_Alarm_Start_M")
   Button "Button_39" at 184,388 size 47x22; TextOff 'Вкл'
      on Click: SetBit("DOx_DB_LED_M1_Alarm_Start_M")
      Appearance <- "DOx_DB_LED_M1_Alarm_Start_M"
   Button "Button_40" at 360,365 size 46x20; TextOff 'Inv'
      on Click: InvertBit("DOx_DB_LED_M1_Alarm_Inverse")
      Appearance <- "DOx_DB_LED_M1_Alarm_Inverse"
   Button "Button_41" at 360,390 size 46x20; TextOff 'Sim'
      on Click: InvertBit("DOx_DB_LED_M1_Alarm_Simulation")
      Appearance <- "DOx_DB_LED_M1_Alarm_Simulation"
   TextField "Text field_15" at 131,425 size 45x22; Text 'Q 0.7'
   TextField "Text field_16" at 176,425 size 120x22; Text 'LED М2 Авария'
   Circle "Circle_15" at 131,448 size 22x22
      Appearance <- "DOx_DB_LED_M2_Alarm_Start_A"
   Circle "Circle_16" at 154,448 size 22x22
      Appearance <- "DOx_DB_LED_M2_Alarm_Q"
   Button "Button_42" at 298,426 size 59x44; TextOff 'Авто'; TextList "Hand"
      on Click: InvertBit("DOx_DB_LED_M2_Alarm_Hand")
      Appearance <- "DOx_DB_LED_M2_Alarm_Hand"
      ProcessValue <- "DOx_DB_LED_M2_Alarm_Hand"
   Button "Button_43" at 240,448 size 49x22; TextOff 'Выкл'
      on Click: ResetBit("DOx_DB_LED_M2_Alarm_Start_M")
   Button "Button_44" at 184,448 size 47x22; TextOff 'Вкл'
      on Click: SetBit("DOx_DB_LED_M2_Alarm_Start_M")
      Appearance <- "DOx_DB_LED_M2_Alarm_Start_M"
   Button "Button_45" at 360,425 size 46x20; TextOff 'Inv'
      on Click: InvertBit("DOx_DB_LED_M2_Alarm_Inverse")
      Appearance <- "DOx_DB_LED_M2_Alarm_Inverse"
   Button "Button_46" at 360,450 size 46x20; TextOff 'Sim'
      on Click: InvertBit("DOx_DB_LED_M2_Alarm_Simulation")
      Appearance <- "DOx_DB_LED_M2_Alarm_Simulation"
   TextField "Text field_17" at 437,10 size 45x22; Text 'Q 1.0'
   TextField "Text field_18" at 482,10 size 120x22; Text 'LED М3 Авария'
   Circle "Circle_17" at 437,33 size 22x22
      Appearance <- "DOx_DB_LED_M3_Alarm_Start_A"
   Circle "Circle_18" at 460,33 size 22x22
      Appearance <- "DOx_DB_LED_M3_Alarm_Q"
   Button "Button_47" at 604,11 size 59x44; TextOff 'Авто'; TextList "Hand"
      on Click: InvertBit("DOx_DB_LED_M3_Alarm_Hand")
      Appearance <- "DOx_DB_LED_M3_Alarm_Hand"
      ProcessValue <- "DOx_DB_LED_M3_Alarm_Hand"
   Button "Button_48" at 546,33 size 49x22; TextOff 'Выкл'
      on Click: ResetBit("DOx_DB_LED_M3_Alarm_Start_M")
   Button "Button_49" at 490,33 size 47x22; TextOff 'Вкл'
      on Click: SetBit("DOx_DB_LED_M3_Alarm_Start_M")
      Appearance <- "DOx_DB_LED_M3_Alarm_Start_M"
   Button "Button_50" at 666,10 size 46x20; TextOff 'Inv'
      on Click: InvertBit("DOx_DB_LED_M3_Alarm_Inverse")
      Appearance <- "DOx_DB_LED_M3_Alarm_Inverse"
   Button "Button_51" at 666,35 size 46x20; TextOff 'Sim'
      on Click: InvertBit("DOx_DB_LED_M3_Alarm_Simulation")
      Appearance <- "DOx_DB_LED_M3_Alarm_Simulation"

screen "About" 800x480, template "Main"
   TextField "Text field_1" at 174,5 size 426x47; Text 'ООО "Водообработка"'
   TextField "Text field_4" at 61,89 size 652x73; Text 'Разработка и поставка оборудования для подготовки реагентов, дозирования, ввода и высокоэффективного перемешивания веществ в непрерывных технологическихх процессах.'
   TextField "Text field_2" at 43,199 size 689x50; Text 'Контактная информация: Адрес: Россия, г. Москва, 111116 ул. Лефортовский вал, д. 7Г, стр. 5'
   TextField "Text field_3" at 238,286 size 299x27; Text 'Телефон: +7 (495) 763-29-73'
   TextField "Text field_5" at 235,313 size 301x27; Text 'http://www.vodoobrabotka.ru'
   GraphicView "Graphic view_1" at 240,358 size 302x96; Picture "logo"

screen "Settings" 800x480, template "Main"
   Button "Button_1" at 7,5 size 96x32; TextOff 'Насосы'; Authorization "Admin"
      on Release: ActivateScreen("Dos", 0); SetTag("settings", 1)
      Appearance <- "settings"
   Button "Button_2" at 7,52 size 96x32; TextOff 'Расход'; Authorization "Admin"
      on Release: ActivateScreen("Flow", 0); SetTag("settings", 2)
      Appearance <- "settings"
   Button "Button_3" at 7,99 size 96x32; TextOff 'Мутность'; Authorization "Admin"
      on Release: ActivateScreen("Trans", 0); SetTag("settings", 3)
      Appearance <- "settings"
   Button "Button_5" at 7,146 size 96x32; TextOff 'DI'; Authorization "Admin"
      on Release: ActivateScreen("DI", 0); SetTag("settings", 4)
      Appearance <- "settings"
   Button "Button_6" at 7,193 size 96x32; TextOff 'DO'; Authorization "Admin"
      on Release: ActivateScreen("DO", 0); SetTag("settings", 5)
      Appearance <- "settings"
   IOField "I/O field_2" at 199,52 size 69x30; FormatPattern 99999
      ProcessValue <- "Time_Today_YEAR"
   IOField "I/O field_1" at 286,52 size 69x30; FormatPattern 999
      ProcessValue <- "Time_Today_MONTH"
   IOField "I/O field_3" at 547,52 size 69x30; FormatPattern 999
      ProcessValue <- "Time_Today_MINUTE"
   IOField "I/O field_4" at 373,52 size 69x30; FormatPattern 999
      ProcessValue <- "Time_Today_DAY"
   IOField "I/O field_5" at 460,52 size 69x30; FormatPattern 999
      ProcessValue <- "Time_Today_HOUR"
   TextField "Text field_4" at 215,29 size 34x23; Text 'год'
   TextField "Text field_1" at 290,29 size 56x23; Text 'месяц'
   TextField "Text field_2" at 386,29 size 45x23; Text 'день'
   TextField "Text field_3" at 477,29 size 33x23; Text 'час'
   TextField "Text field_5" at 547,29 size 68x23; Text 'минуты'
   IOField "I/O field_6" at 200,116 size 69x30; FormatPattern 99999
      ProcessValue <- "Time_Year"
   IOField "I/O field_7" at 287,116 size 69x30; FormatPattern 99999
      ProcessValue <- "Time_Month"
   IOField "I/O field_8" at 548,116 size 69x30; FormatPattern 99999
      ProcessValue <- "Time_Minutes"
   IOField "I/O field_9" at 374,116 size 69x30; FormatPattern 99999
      ProcessValue <- "Time_Day"
   IOField "I/O field_10" at 461,116 size 69x30; FormatPattern 99999
      ProcessValue <- "Time_Hour"
   TextField "Text field_6" at 216,93 size 34x23; Text 'год'
   TextField "Text field_7" at 291,93 size 56x23; Text 'месяц'
   TextField "Text field_8" at 387,93 size 45x23; Text 'день'
   TextField "Text field_9" at 478,93 size 33x23; Text 'час'
   TextField "Text field_10" at 548,93 size 68x23; Text 'минуты'
   Button "Button_4" at 526,170 size 90x22; TextOff 'Сохранить'; TextList "Hand"
      on Click: SetBit("Time_Save")
      ProcessValue <- "Motors_DB_M1_CMD_Hand"

